(* Logix 5000 project; controller MV vendor 1 type 14 code 217 rev 31.11; software revision 31.00 *) (continued)
   MC_CH1_Log_ID : DINT := 56;
   MC_CH1_OneShot : BOOL;
   MC_CH1_PR1 : PlantItem := (CW := 2#0000_0000_0000_0000_0000_0000_0001_0000, CheckTime := 8, CheckTimer := 8);   // CH1_PR1
   MC_CH1_PR1_ALARM : ALARM_DIGITAL;
   MC_CH1_PR1_C : ALIAS FOR RIO_Rack_2:6:I.Data.6;
   MC_CH1_PR1_DR : ALIAS FOR RIO_Rack_2:5:O.Data.18;
   MC_CH1_PR1_O : ALIAS FOR RIO_Rack_2:6:I.Data.2;
   MC_CH1_PTX_AI : PlantItem := (CW := 2#0000_0000_0000_0000_1000_0000_0000_0000, CheckTime := 15, CheckTimer := 15, Scaled := 55.846878, RawInput := 9957.0);   // CH1_PTX
   MC_CH1_PTX_AI_RawInput : ALIAS FOR RIO_Rack_2:1:I.Ch6Data;   // Real Analog Input , Do Not Use In Code
   MC_CH1_R1 : PlantItem := (CW := 2#0000_0000_0000_0000_0000_0000_0011_0000, CheckTime := 20, CheckTimer := 20);   // CH1_R1
   MC_CH1_R1_ALARM : ALARM_DIGITAL;
   MC_CH1_R1_C : ALIAS FOR RIO_Rack_2:4:I.Data.4;
   MC_CH1_R1_DR : ALIAS FOR RIO_Rack_2:5:O.Data.0;
   MC_CH1_R1_O : ALIAS FOR RIO_Rack_2:4:I.Data.0;
   MC_CH1_R1R : PlantItem := (CW := 2#0000_0000_0000_0000_0000_0000_0001_0000, CheckTime := 20, CheckTimer := 20);   // CH1_R1R
   MC_CH1_R1R_ALARM : ALARM_DIGITAL;
   MC_CH1_R1R_C : ALIAS FOR RIO_Rack_2:4:I.Data.14;
   MC_CH1_R1R_DR : ALIAS FOR RIO_Rack_2:5:O.Data.6;
   MC_CH1_R1R_O : ALIAS FOR RIO_Rack_2:4:I.Data.10;
   MC_CH1_R2 : PlantItem := (CW := 2#0000_0000_0000_0000_0000_0000_0001_0000, CheckTime := 20, CheckTimer := 20);   // CH1_R2
   MC_CH1_R2_ALARM : ALARM_DIGITAL;
   MC_CH1_R2_C : ALIAS FOR RIO_Rack_2:4:I.Data.5;
   MC_CH1_R2_DR : ALIAS FOR RIO_Rack_2:5:O.Data.1;
   MC_CH1_R2_O : ALIAS FOR RIO_Rack_2:4:I.Data.1;
   MC_CH1_R2R : PlantItem := (CW := 2#0000_0000_0000_0000_0000_0000_0001_0000, CheckTime := 20, CheckTimer := 20);   // CH1_R2R
   MC_CH1_R2R_ALARM : ALARM_DIGITAL;
   MC_CH1_R2R_C : ALIAS FOR RIO_Rack_2:4:I.Data.15;
   MC_CH1_R2R_DR : ALIAS FOR RIO_Rack_2:5:O.Data.7;
   MC_CH1_R2R_O : ALIAS FOR RIO_Rack_2:4:I.Data.11;
   MC_CH1_R3 : PlantItem := (CW := 2#0000_0000_0000_0000_0000_0000_0001_0000, CheckTime := 20, CheckTimer := 20);   // CH1_R3
   MC_CH1_R3_ALARM : ALARM_DIGITAL;
   MC_CH1_R3_C : ALIAS FOR RIO_Rack_2:4:I.Data.6;
   MC_CH1_R3_DR : ALIAS FOR RIO_Rack_2:5:O.Data.2;
   MC_CH1_R3_O : ALIAS FOR RIO_Rack_2:4:I.Data.2;
   MC_CH1_R3R : PlantItem := (CW := 2#0000_0000_0000_0000_0000_0000_0001_0000, CheckTime := 20, CheckTimer := 20);   // CH1_R3R
   MC_CH1_R3R_ALARM : ALARM_DIGITAL;
   MC_CH1_R3R_C : ALIAS FOR RIO_Rack_2:4:I.Data.20;
   MC_CH1_R3R_DR : ALIAS FOR RIO_Rack_2:5:O.Data.8;
   MC_CH1_R3R_O : ALIAS FOR RIO_Rack_2:4:I.Data.16;
   MC_CH1_R4 : PlantItem := (CW := 2#0000_0000_0000_0000_0000_0000_0001_0000, CheckTime := 20, CheckTimer := 20);   // CH1_R4
   MC_CH1_R4_ALARM : ALARM_DIGITAL;
   MC_CH1_R4_C : ALIAS FOR RIO_Rack_2:4:I.Data.7;
   MC_CH1_R4_DR : ALIAS FOR RIO_Rack_2:5:O.Data.3;
   MC_CH1_R4_O : ALIAS FOR RIO_Rack_2:4:I.Data.3;
   MC_CH1_R4R : PlantItem := (CW := 2#0000_0000_0000_0000_0000_0000_0001_0000, CheckTime := 20, CheckTimer := 20);   // CH1_R4R
   MC_CH1_R4R_ALARM : ALARM_DIGITAL;
   MC_CH1_R4R_C : ALIAS FOR RIO_Rack_2:4:I.Data.21;
   MC_CH1_R4R_DR : ALIAS FOR RIO_Rack_2:5:O.Data.9;
   MC_CH1_R4R_O : ALIAS FOR RIO_Rack_2:4:I.Data.17;
   MC_CH1_R5 : PlantItem := (CW := 2#0000_0000_0000_0000_0000_0000_0001_0000, CheckTime := 20, CheckTimer := 20);   // CH1_R5
   MC_CH1_R5_ALARM : ALARM_DIGITAL;
   MC_CH1_R5_C : ALIAS FOR RIO_Rack_2:4:I.Data.12;
   MC_CH1_R5_DR : ALIAS FOR RIO_Rack_2:5:O.Data.4;
   MC_CH1_R5_O : ALIAS FOR RIO_Rack_2:4:I.Data.8;
   MC_CH1_R5R : PlantItem := (CW := 2#0000_0000_0000_0000_0000_0000_0001_0000, CheckTime := 20, CheckTimer := 20);   // CH1_R5R
   MC_CH1_R5R_ALARM : ALARM_DIGITAL;
   MC_CH1_R5R_C : ALIAS FOR RIO_Rack_2:4:I.Data.22;
   MC_CH1_R5R_DR : ALIAS FOR RIO_Rack_2:5:O.Data.10;
   MC_CH1_R5R_O : ALIAS FOR RIO_Rack_2:4:I.Data.18;
   MC_CH1_R6 : PlantItem := (CW := 2#0000_0000_0000_0000_0000_0000_1000_1011, CheckTime := 20, CheckTimer := 20, DriveBits := 1);   // CH1_R6
   MC_CH1_R6_ALARM : ALARM_DIGITAL;
   MC_CH1_R6_C : ALIAS FOR RIO_Rack_2:4:I.Data.13;
   MC_CH1_R6_DR : ALIAS FOR RIO_Rack_2:5:O.Data.5;
   MC_CH1_R6_O : ALIAS FOR RIO_Rack_2:4:I.Data.9;
   MC_CH1_R6R : PlantItem := (CW := 2#0000_0000_0000_0000_0000_0000_1000_1011, CheckTime := 20, CheckTimer := 20, DriveBits := 1);   // CH1_R6R
   MC_CH1_R6R_ALARM : ALARM_DIGITAL;
   MC_CH1_R6R_C : ALIAS FOR RIO_Rack_2:4:I.Data.23;
   MC_CH1_R6R_DR : ALIAS FOR RIO_Rack_2:5:O.Data.11;
   MC_CH1_R6R_O : ALIAS FOR RIO_Rack_2:4:I.Data.19;
   MC_CH1_RESET : ALIAS FOR MC_N100[30].0;   // CH1 reset flag
   MC_CH1_RESTART : ALIAS FOR MC_N100[35];   // CH1 restart step
   MC_CH1_RETURN : ALIAS FOR MC_N100[32].7;   // CH1 open return route flag
   MC_CH1_RP_OFF : ALIAS FOR MC_N100[32].2;   // CH1 enable return pump off delay timer
   MC_CH1_RP_ON : ALIAS FOR MC_N100[32].1;   // CH1 enable return pump on delay timer
   MC_CH1_RPUMP : ALIAS FOR MC_N100[32].4;   // CH1 run return pump flag
   MC_CH1_RR : PlantItem := (CW := 2#0000_0000_0000_0000_0000_0000_0001_0000, CheckTime := 20, CheckTimer := 20);   // CH1_RR
   MC_CH1_RR_ALARM : ALARM_DIGITAL;
   MC_CH1_RR_C : ALIAS FOR RIO_Rack_2:4:I.Data.29;
   MC_CH1_RR_DR : ALIAS FOR RIO_Rack_2:5:O.Data.13;
   MC_CH1_RR_O : ALIAS FOR RIO_Rack_2:4:I.Data.25;
   MC_CH1_RTNFLOW : ALIAS FOR MC_N100[18].0;   // CH1 Is Return Flow flag
   MC_CH1_SaveCIPReport_now : DINT;
   MC_CH1_SaveCIPReport_now_done : DINT := -1;
   MC_CH1_STATUS : ALIAS FOR MC_N100[0];   // CH1 status 0: Unavailable; 1: Idle; 2: Running; 3: Stopped; 4: Faulted
   MC_CH1_SUBSTEP : ALIAS FOR MC_N100[17];   // CH1 current substep
   MC_CH1_SUPPLY : ALIAS FOR MC_N100[32].3;   // CH1 open supply route flag
   MC_CH1_T105_2_ACC : DINT := 86383;
   MC_CH1_TIMING : ALIAS FOR MC_N100[30].3;   // CH1 run current cycle timer
   MC_CH1_TODET : ALIAS FOR MC_N100[18].2;   // CH1 return postrinse to detergent tank
   MC_CH2_ACTIVE : ALIAS FOR MC_N120[30].1;   // CH2 active flag
   MC_CH2_CIP_BYPASS_Conditions : BOOL;
   MC_CH2_CIP_BYPASS_DrainConditions : BOOL;
   MC_CH2_CIP_Messages : STRING[20];   // CH2 CIP Scada Messages
        [4]   // Channel 2 CIP Completion Clock Time
        [0]   // Channel 2 CIP Program Text for Scada
        [1]   // Channel2 CIP Cycle Text for Scada
        [2]   // Channel 2 CIP Time Left Text for Scada
        [3]   // Channel 2 CIP Down Time Text for Scada
   MC_CH2_CIP_Misc : DINT[20];
   MC_CH2_CIP_MiscReal : REAL[20];
   MC_CH2_CIP_YST_Scb_Bypass : BOOL;
   MC_CH2_CSTEP : ALIAS FOR MC_N120[34];   // CH2 command processor current step
   MC_CH2_CTX2_AI : PlantItem := (CW := 2#0000_0000_0000_0000_1000_0000_0000_0000, CheckTime := 15, CheckTimer := 15, Scaled := 0.00875, RawInput := 4014.0);   // CH2_CTX2
   MC_CH2_CTX2_AI_RawInput : ALIAS FOR RIO_Rack_2:1:I.Ch3Data;   // Real Analog Input , Do Not Use In Code
   MC_CH2_CYCDONE : ALIAS FOR MC_T125[2].DN;   // CH2 current cycle complete
   MC_CH2_CYCLE : ALIAS FOR MC_N120[1];   // CH2 current CIP cycle
   MC_CH2_Delay_For_Data : TIMER := (PRE := 2000);
   MC_CH2_DETRTN : ALIAS FOR MC_N120[18].1;   // CH2 Is Detergent Return flag
   MC_CH2_DONE : ALIAS FOR MC_N120[30].4;   // CH2 cycle complete flag
   MC_CH2_DR1 : PlantItem := (CW := 2#0000_0000_0000_0000_0000_0000_0001_0000, CheckTime := 8, CheckTimer := 8);   // CH2_DR1
   MC_CH2_DR1_ALARM : ALARM_DIGITAL;
   MC_CH2_DR1_C : ALIAS FOR RIO_Rack_2:7:I.Data.6;
   MC_CH2_DR1_DR : ALIAS FOR RIO_Rack_2:8:O.Data.2;
   MC_CH2_DR1_O : ALIAS FOR RIO_Rack_2:7:I.Data.2;
   MC_CH2_DR2 : PlantItem := (CW := 2#0000_0000_0000_0000_0000_0000_0001_0000, CheckTime := 8, CheckTimer := 8);   // CH2_DR2
   MC_CH2_DR2_ALARM : ALARM_DIGITAL;
   MC_CH2_DR2_C : ALIAS FOR RIO_Rack_2:7:I.Data.7;
   MC_CH2_DR2_DR : ALIAS FOR RIO_Rack_2:8:O.Data.3;
   MC_CH2_DR2_O : ALIAS FOR RIO_Rack_2:7:I.Data.3;
   MC_CH2_DRAIN : PlantItem := (CW := 2#0000_0000_0000_0000_0000_0000_0001_0000, CheckTime := 8, CheckTimer := 8);   // CH2_DRAIN
   MC_CH2_DRAIN_ALARM : ALARM_DIGITAL;
   MC_CH2_DRAIN_C : ALIAS FOR RIO_Rack_2:7:I.Data.4;
   MC_CH2_DRAIN_CLOSE : BOOL;
   MC_CH2_DRAIN_DR : ALIAS FOR RIO_Rack_2:8:O.Data.0;
   MC_CH2_DRAIN_O : ALIAS FOR RIO_Rack_2:7:I.Data.0;
   MC_CH2_DT : ALIAS FOR MC_N120[10];   // CH2 detergent tank to use (1 or 2)
   MC_CH2_DT1 : PlantItem := (CW := 2#0000_0000_0000_0000_0000_0000_0001_0000, CheckTime := 8, CheckTimer := 8);   // CH2_DT1
   MC_CH2_DT1_ALARM : ALARM_DIGITAL;
   MC_CH2_DT1_C : ALIAS FOR RIO_Rack_2:7:I.Data.12;
   MC_CH2_DT1_DR : ALIAS FOR RIO_Rack_2:8:O.Data.4;
   MC_CH2_DT1_O : ALIAS FOR RIO_Rack_2:7:I.Data.8;
   MC_CH2_DT2 : PlantItem := (CW := 2#0000_0000_0000_0000_0000_0000_0001_0000, CheckTime := 12, CheckTimer := 12);   // CH2_DT2
   MC_CH2_DT2_ALARM : ALARM_DIGITAL;
   MC_CH2_DT2_C : ALIAS FOR RIO_Rack_2:7:I.Data.13;
   MC_CH2_DT2_DR : ALIAS FOR RIO_Rack_2:8:O.Data.5;
   MC_CH2_DT2_O : ALIAS FOR RIO_Rack_2:7:I.Data.9;
   MC_CH2_EVENT : ALIAS FOR MC_N120[23];   // CH2 event register
   MC_CH2_EXTEND : ALIAS FOR MC_N120[30].5;   // CH2 extend cycle flag
   MC_CH2_FAULT : ALIAS FOR MC_N120[20];   // CH2 fault register
   MC_CH2_FM_AI : PlantItem := (CW := 2#0000_0000_0000_0000_1000_0000_0000_0000, CheckTime := 15, CheckTimer := 15, Scaled := 1.0, RawInput := 4032.0);   // CH2_FM
   MC_CH2_FM_AI_RawInput : ALIAS FOR RIO_Rack_2:1:I.Ch5Data;   // Real Analog Input , Do Not Use In Code
   MC_CH2_FVBypass_Flush_ALARM : ALARM_DIGITAL;
   MC_CH2_FVBYPASS_H2O_Flush : BOOL;
   MC_CH2_ISLINE : ALIAS FOR MC_N122[13].0;   // CH2 Is Line Clean flag
   MC_CH2_LF1 : PlantItem := (CW := 2#0000_0000_0000_0000_0000_0000_0001_0000, CheckTime := 8, CheckTimer := 8);   // CH2_LF1
   MC_CH2_LF1_ALARM : ALARM_DIGITAL;
   MC_CH2_LF1_C : ALIAS FOR RIO_Rack_2:7:I.Data.15;
   MC_CH2_LF1_DR : ALIAS FOR RIO_Rack_2:8:O.Data.7;
   MC_CH2_LF1_O : ALIAS FOR RIO_Rack_2:7:I.Data.11;
   MC_CH2_Log_ID : DINT := 57;
   MC_CH2_OneShot : BOOL;
   MC_CH2_PR1 : PlantItem := (CW := 2#0000_0000_0000_0000_0000_0000_0001_0000, CheckTime := 8, CheckTimer := 8);   // CH2_PR1
   MC_CH2_PR1_ALARM : ALARM_DIGITAL;
   MC_CH2_PR1_C : ALIAS FOR RIO_Rack_2:7:I.Data.14;
   MC_CH2_PR1_DR : ALIAS FOR RIO_Rack_2:8:O.Data.6;
   MC_CH2_PR1_O : ALIAS FOR RIO_Rack_2:7:I.Data.10;
   MC_CH2_PTX_AI : PlantItem := (CW := 2#0000_0000_0000_0000_1000_0000_0000_0000, CheckTime := 15, CheckTimer := 15, Scaled := 8.446876, RawInput := 4901.0);   // CH2_PTX
   MC_CH2_PTX_AI_RawInput : ALIAS FOR RIO_Rack_2:1:I.Ch7Data;   // Real Analog Input , Do Not Use In Code
   MC_CH2_R1 : PlantItem := (CW := 2#0000_0000_0000_0000_0000_0000_0001_0000, CheckTime := 8, CheckTimer := 8);   // CH2_R1
   MC_CH2_R1_ALARM : ALARM_DIGITAL;
   MC_CH2_R1_C : ALIAS FOR RIO_Rack_2:6:I.Data.12;
   MC_CH2_R1_DR : ALIAS FOR RIO_Rack_2:5:O.Data.20;
   MC_CH2_R1_O : ALIAS FOR RIO_Rack_2:6:I.Data.8;
   MC_CH2_R1R : PlantItem := (CW := 2#0000_0000_0000_0000_0000_0000_0001_0000, CheckTime := 8, CheckTimer := 8);   // CH2_R1R
   MC_CH2_R1R_ALARM : ALARM_DIGITAL;
   MC_CH2_R1R_C : ALIAS FOR RIO_Rack_2:6:I.Data.22;
   MC_CH2_R1R_DR : ALIAS FOR RIO_Rack_2:5:O.Data.26;
   MC_CH2_R1R_O : ALIAS FOR RIO_Rack_2:6:I.Data.18;
   MC_CH2_R2 : PlantItem := (CW := 2#0000_0000_0000_0000_0000_0000_0001_0000, CheckTime := 8, CheckTimer := 8);   // CH2_R2
   MC_CH2_R2_ALARM : ALARM_DIGITAL;
   MC_CH2_R2_C : ALIAS FOR RIO_Rack_2:6:I.Data.13;
   MC_CH2_R2_DR : ALIAS FOR RIO_Rack_2:5:O.Data.21;
   MC_CH2_R2_O : ALIAS FOR RIO_Rack_2:6:I.Data.9;
   MC_CH2_R2R : PlantItem := (CW := 2#0000_0000_0000_0000_0000_0000_0001_0000, CheckTime := 8, CheckTimer := 8);   // CH2_R2R
   MC_CH2_R2R_ALARM : ALARM_DIGITAL;
   MC_CH2_R2R_C : ALIAS FOR RIO_Rack_2:6:I.Data.23;
   MC_CH2_R2R_DR : ALIAS FOR RIO_Rack_2:5:O.Data.27;
   MC_CH2_R2R_O : ALIAS FOR RIO_Rack_2:6:I.Data.19;
   MC_CH2_R3 : PlantItem := (CW := 2#0000_0000_0000_0000_0000_0000_0001_0000, CheckTime := 8, CheckTimer := 8);   // CH2_R3
   MC_CH2_R3_ALARM : ALARM_DIGITAL;
   MC_CH2_R3_C : ALIAS FOR RIO_Rack_2:6:I.Data.14;
   MC_CH2_R3_DR : ALIAS FOR RIO_Rack_2:5:O.Data.22;
   MC_CH2_R3_O : ALIAS FOR RIO_Rack_2:6:I.Data.10;
   MC_CH2_R3R : PlantItem := (CW := 2#0000_0000_0000_0000_0000_0000_0001_0000, CheckTime := 8, CheckTimer := 8);   // CH2_R3R
   MC_CH2_R3R_ALARM : ALARM_DIGITAL;
   MC_CH2_R3R_C : ALIAS FOR RIO_Rack_2:6:I.Data.28;
   MC_CH2_R3R_DR : ALIAS FOR RIO_Rack_2:5:O.Data.28;
   MC_CH2_R3R_O : ALIAS FOR RIO_Rack_2:6:I.Data.24;
   MC_CH2_R4 : PlantItem := (CW := 2#0000_0000_0000_0000_0000_0000_0001_0000, CheckTime := 8, CheckTimer := 8);   // CH2_R4
   MC_CH2_R4_ALARM : ALARM_DIGITAL;
   MC_CH2_R4_C : ALIAS FOR RIO_Rack_2:6:I.Data.15;
   MC_CH2_R4_DR : ALIAS FOR RIO_Rack_2:5:O.Data.23;
   MC_CH2_R4_O : ALIAS FOR RIO_Rack_2:6:I.Data.11;
   MC_CH2_R4R : PlantItem := (CW := 2#0000_0000_0000_0000_0000_0000_0001_0000, CheckTime := 8, CheckTimer := 8);   // CH2_R4R
   MC_CH2_R4R_ALARM : ALARM_DIGITAL;
   MC_CH2_R4R_C : ALIAS FOR RIO_Rack_2:6:I.Data.29;
   MC_CH2_R4R_DR : ALIAS FOR RIO_Rack_2:5:O.Data.29;
   MC_CH2_R4R_O : ALIAS FOR RIO_Rack_2:6:I.Data.25;
   MC_CH2_R5 : PlantItem := (CW := 2#0000_0000_0000_0000_0000_0000_0001_0000, CheckTime := 8, CheckTimer := 8);   // CH2_R5
   MC_CH2_R5_ALARM : ALARM_DIGITAL;
   MC_CH2_R5_C : ALIAS FOR RIO_Rack_2:6:I.Data.20;
   MC_CH2_R5_DR : ALIAS FOR RIO_Rack_2:5:O.Data.24;
   MC_CH2_R5_O : ALIAS FOR RIO_Rack_2:6:I.Data.16;
   MC_CH2_R5R : PlantItem := (CW := 2#0000_0000_0000_0000_0000_0000_0001_0000, CheckTime := 8, CheckTimer := 8);   // CH2_R5R
   MC_CH2_R5R_ALARM : ALARM_DIGITAL;
   MC_CH2_R5R_C : ALIAS FOR RIO_Rack_2:6:I.Data.30;
   MC_CH2_R5R_DR : ALIAS FOR RIO_Rack_2:5:O.Data.30;
   MC_CH2_R5R_O : ALIAS FOR RIO_Rack_2:6:I.Data.26;
   MC_CH2_R6 : PlantItem := (CW := 2#0000_0000_0000_0000_0000_0001_0001_0000, CheckTime := 8, CheckTimer := 8);   // CH2_R6
   MC_CH2_R6_ALARM : ALARM_DIGITAL;
   MC_CH2_R6_C : ALIAS FOR RIO_Rack_2:6:I.Data.21;
   MC_CH2_R6_DR : ALIAS FOR RIO_Rack_2:5:O.Data.25;
   MC_CH2_R6_O : ALIAS FOR RIO_Rack_2:6:I.Data.17;
   MC_CH2_R6R : PlantItem := (CW := 2#0000_0000_0000_0000_0000_0000_0001_0000, CheckTime := 8, CheckTimer := 8);   // CH2_R6R
   MC_CH2_R6R_ALARM : ALARM_DIGITAL;
   MC_CH2_R6R_C : ALIAS FOR RIO_Rack_2:6:I.Data.31;
   MC_CH2_R6R_DR : ALIAS FOR RIO_Rack_2:5:O.Data.31;
   MC_CH2_R6R_O : ALIAS FOR RIO_Rack_2:6:I.Data.27;
   MC_CH2_RESET : ALIAS FOR MC_N120[30].0;   // CH2 reset flag
   MC_CH2_RESTART : ALIAS FOR MC_N120[35];   // CH2 restart step
   MC_CH2_RETURN : ALIAS FOR MC_N120[32].7;   // CH2 open return route flag
   MC_CH2_RP_ON : ALIAS FOR MC_N120[32].1;   // CH2 enable return pump on delay timer
   MC_CH2_RPUMP : ALIAS FOR MC_N120[32].4;   // CH2 run return pump flag
   MC_CH2_RR : PlantItem := (CW := 2#0000_0000_0000_0000_0000_0000_0001_0000, CheckTime := 8, CheckTimer := 8);   // CH2_RR
   MC_CH2_RR_ALARM : ALARM_DIGITAL;
   MC_CH2_RR_C : ALIAS FOR RIO_Rack_2:7:I.Data.5;
   MC_CH2_RR_DR : ALIAS FOR RIO_Rack_2:8:O.Data.1;
   MC_CH2_RR_O : ALIAS FOR RIO_Rack_2:7:I.Data.1;
   MC_CH2_RTNFLOW : ALIAS FOR MC_N120[18].0;   // CH2 return flow on debounce timer
   MC_CH2_SaveCIPReport_now : DINT;
   MC_CH2_SaveCIPReport_now_done : DINT := -1;
   MC_CH2_STATUS : ALIAS FOR MC_N120[0];   // CH2 status 0: Unavailable; 1: Idle; 2: Running; 3: Stopped; 4: Faulted
   MC_CH2_SUBSTEP : ALIAS FOR MC_N120[17];   // CH2 current substep
   MC_CH2_SUPPLY : ALIAS FOR MC_N120[32].3;   // CH2 open supply route flag
   MC_CH2_T125_2_ACC : DINT := 90000;
   MC_CH2_TIMING : ALIAS FOR MC_N120[30].3;   // CH2 run current cycle timer
   MC_CH2_TODET : ALIAS FOR MC_N120[18].2;   // CH2 return postrinse to detergent tank
   MC_CH2_TURBID_High : BOOL;
   MC_Channel1_Channel_1_event : STRING;
   MC_Channel1_Channel_1_event_prefix : STRING;
   MC_Channel1_Channel_2_event : STRING;
   MC_Channel1_Channel_2_event_prefix : STRING;
   MC_CIP_AV01 : PlantItem := (CW := 2#0000_0000_0000_0000_0000_0000_1000_1011, CheckTime := 8, CheckTimer := 8, DriveBits := 1);   // CIP_AV01
   MC_CIP_AV01_ALARM : ALARM_DIGITAL;
   MC_CIP_AV01_C : ALIAS FOR RIO_Rack_2:9:I.Data.23;
   MC_CIP_AV01_DR : ALIAS FOR CIP_AV01_DUMMY_DR;
   MC_CIP_AV01_O : ALIAS FOR RIO_Rack_2:9:I.Data.19;
   MC_CIP_AV02 : PlantItem := (CW := 2#0000_0000_0000_0000_0000_0000_0001_0000, CheckTime := 8, CheckTimer := 8);   // CIP_AV02
   MC_CIP_AV02_ALARM : ALARM_DIGITAL;
   MC_CIP_AV02_C : ALIAS FOR RIO_Rack_2:9:I.Data.28;
   MC_CIP_AV02_DR : ALIAS FOR RIO_Rack_2:8:O.Data.27;   // Used As Output Share Item Rung 20
   MC_CIP_AV02_O : ALIAS FOR RIO_Rack_2:9:I.Data.24;
   MC_CIP_AV05 : PlantItem := (CW := 2#0000_0000_0000_0000_0000_0000_1000_1011, CheckTime := 8, CheckTimer := 8, DriveBits := 1);   // CIP_AV05
   MC_CIP_AV05_ALARM : ALARM_DIGITAL;
   MC_CIP_AV05_C : ALIAS FOR RIO_Rack_2:9:I.Data.29;
   MC_CIP_AV05_DR : ALIAS FOR CIP_AV05_DUMMY_DR;
   MC_CIP_AV05_O : ALIAS FOR RIO_Rack_2:9:I.Data.25;
   MC_CIP_AV06 : PlantItem := (CW := 2#0000_0000_0000_0000_0000_0000_0001_0000, CheckTime := 8, CheckTimer := 8);   // CIP_AV06
   MC_CIP_AV06_ALARM : ALARM_DIGITAL;
   MC_CIP_AV06_C : ALIAS FOR RIO_Rack_2:9:I.Data.30;
   MC_CIP_AV06_DR : ALIAS FOR RIO_Rack_2:8:O.Data.28;
   MC_CIP_AV06_O : ALIAS FOR RIO_Rack_2:9:I.Data.26;
   MC_CIP_AV07 : PlantItem := (CW := 2#0000_0000_0000_0000_0000_0000_1000_1011, CheckTime := 8, CheckTimer := 8, DriveBits := 1);   // CIP_AV07
   MC_CIP_AV07_ALARM : ALARM_DIGITAL;
   MC_CIP_AV07_C : ALIAS FOR RIO_Rack_2:9:I.Data.31;
   MC_CIP_AV07_DR : ALIAS FOR CIP_AV07_DUMMY_DR;
   MC_CIP_AV07_O : ALIAS FOR RIO_Rack_2:9:I.Data.27;
   MC_CIP_AV08 : PlantItem := (CW := 2#0000_0000_0000_0000_0000_0000_0001_0000, CheckTime := 8, CheckTimer := 8);   // CIP_AV08
   MC_CIP_AV08_ALARM : ALARM_DIGITAL;
   MC_CIP_AV08_C : ALIAS FOR RIO_Rack_2:11:I.Data.20;
   MC_CIP_AV08_DR : ALIAS FOR RIO_Rack_2:8:O.Data.29;
   MC_CIP_AV08_O : ALIAS FOR RIO_Rack_2:11:I.Data.24;
   MC_CIP_AV09 : PlantItem := (CW := 2#0000_0000_0000_0000_0000_0000_1000_1011, CheckTime := 8, CheckTimer := 8, DriveBits := 1);   // CIP_AV09
   MC_CIP_AV09_ALARM : ALARM_DIGITAL;
   MC_CIP_AV09_C : ALIAS FOR RIO_Rack_2:11:I.Data.21;
   MC_CIP_AV09_DR : ALIAS FOR CIP_AV09_DUMMY_DR;
   MC_CIP_AV09_O : ALIAS FOR RIO_Rack_2:11:I.Data.25;
   MC_CIP_AV10 : PlantItem := (CW := 2#0000_0000_0000_0000_0000_0000_0001_0000, CheckTime := 8, CheckTimer := 8);   // CIP_AV10
   MC_CIP_AV10_ALARM : ALARM_DIGITAL;
   MC_CIP_AV10_C : ALIAS FOR RIO_Rack_2:11:I.Data.22;
   MC_CIP_AV10_DR : ALIAS FOR RIO_Rack_2:8:O.Data.30;
   MC_CIP_AV10_O : ALIAS FOR RIO_Rack_2:11:I.Data.26;
   MC_CIP_CH2_String_OK : BOOL;
   MC_CIP_CH2_Strings_HopRinse : STRING[30] := ([0] := 'FV', [1] := 'YSV', [2] := 'YPV', [3] := 'YCV', [4] := 'Yeast Pitch Main', [5] := 'Yeast Slurry Tank', [6] := 'Gales Yeast Main', [7] := 'YSV1 Reseeding Line', [8] := 'Filtrate Tank', [9] := 'Yeast Main FVs1 to 17 Short', [10] := 'Yeast Main FVs1 to 17 Long', [11] := 'Yeast Main FVs18 to 25 Short', [12] := 'Yeast Main FVs18 to 25 Long', [13] := 'Yeast Room and Pump', [14] := 'FVs 26 to 31 Yeast Main Short', [15] := 'FVs 26 to 31 Yeast Main Long', [16] := ' Normal Clean', [17] := ' Hop Rinse', [18] := ' Hop Normal clean 3 pre rinses', [19] := ' Initial rinse', [20] := ' Pre-CIP Initial Rinse', [21] := ' Normal', [22] := 'Cold Water Rinse');
   MC_CIP_Default_Messages : STRING[20] := ([1] := 'Scavenge ', [2] := 'Pre Rinse ', [3] := 'Detergent ', [4] := 'Post Rinse ', [5] := ' of ', [6] := ':', [7] := '0', [17] := '3', [18] := '16', [19] := '1');
        [5]   // cycle of with spaces
        [6]   // colon : for time
        [17]   // Temp Working Area
        [18]   // Temp Working Area
        [0]   // temp area to build
        [19]   // Temp Working Area
        [7]   // leading 'zero'
   MC_CIP_EFFTank_Full : BOOL;
   MC_CIP_EFFTank_Full_Spt : DINT := 50000;
   MC_CIP_EFFTank_Start_Lvl_Ok : BOOL := 1;
   MC_CIP_RV : PlantItem := (CW := 2#0000_0000_0000_0000_0000_0001_0000_0000, CheckTime := 15, CheckTimer := 15);   // CIP_RV
   MC_CIP_RV_ALARM : ALARM_DIGITAL;
   MC_CIP_RV_C : ALIAS FOR RIO_Rack_2:9:I.Data.21;
   MC_CIP_RV_DR : ALIAS FOR RIO_Rack_2:8:O.Data.26;
   MC_CIP_RV_O : ALIAS FOR RIO_Rack_2:9:I.Data.17;
   MC_CIP_String_Result : DINT;
   MC_CIP_temp : INT;
   MC_CLOCK_system_set : BOOL;
   MC_COMMS_FROM_BLUNGER : MESSAGE;
        MessageParameters(ServiceCode := 16#0fa2, LocalElement := MC_N114[0], ...)
   mc_comms_from_brewhouse : MESSAGE;
        MessageParameters(ServiceCode := 16#004c, LocalElement := BH_Draindown_ON, ...)
   mc_comms_from_brewhouse_timer : TIMER := (PRE := 6000, ACC := 1632, EN := 1, TT := 1);
   MC_COMMS_FROM_FV_ROUTING_PLC : MESSAGE;
        MessageParameters(ServiceCode := 16#004c, LocalElement := MC_N112[0], ...)
   MC_COMMS_FROM_MV_ROUTING_PLC : MESSAGE;
        MessageParameters(ServiceCode := 16#004c, LocalElement := MC_N113[0], ...)
   mc_comms_to_blunger : MESSAGE;
        MessageParameters(ServiceCode := 16#0faa, LocalElement := MC_N114[100], ...)
   mc_comms_to_blunger_timer : TIMER := (PRE := 6000, ACC := 631, EN := 1, TT := 1);
   mc_comms_to_fv_route : MESSAGE;
        MessageParameters(ServiceCode := 16#0faa, LocalElement := MC_N112[100], ...)
   mc_comms_to_fv_route_timer : TIMER := (PRE := 6000, ACC := 2121, EN := 1, TT := 1);
   mc_comms_to_mv_route : MESSAGE;
        MessageParameters(ServiceCode := 16#0faa, LocalElement := MC_N113[100], ...)
   mc_comms_to_mv_route_timer : TIMER := (PRE := 6000, ACC := 629, EN := 1, TT := 1);
   MC_copy_how_many : DINT;
   MC_CopyOfCh1Route : DINT := 1032;
   MC_CopyOfCh2Route : DINT := 7;
   MC_CP1 : PlantItem := (CheckTime := 8);   // CP1
   MC_CP1_RawOutput : ALIAS FOR RIO_Rack_2:10:O.Data.14;   // MC_CP1
   MC_CTX_001_AI : PlantItem := (CW := 2#0000_0000_0000_0000_1100_0000_0000_0000, CheckTime := 15, CheckTimer := 15, Scaled := 2.2806249, RawInput := 7649.0);   // CTX_001
   MC_CTX_001_AI_RawInput : ALIAS FOR RIO_Rack_2:1:I.Ch0Data;   // Real Analog Input , Do Not Use In Code
   MC_CTX_002_AI : PlantItem := (CW := 2#0000_0000_0000_0000_1000_0000_0000_0000, CheckTime := 15, CheckTimer := 15, Scaled := 2.170625, RawInput := 7473.0);   // CTX_002
   MC_CTX_002_AI_RawInput : ALIAS FOR RIO_Rack_2:1:I.Ch1Data;   // Real Analog Input , Do Not Use In Code
   MC_data_file_address : DINT := 80;
   MC_data_file_value_to_move : DINT := 18;
   MC_Delphi_I : DINT[60] := ([38] := 29712, [39] := 33151);
   MC_DetTank1_Service_event : STRING;
   MC_DetTank1_Service_event_prefix : STRING;
   MC_DetTank2_Service_event : STRING;
   MC_DetTank2_Service_event_prefix : STRING;
   MC_DT1_CP1 : ALIAS FOR MC_N80[18].8;   // DT1 service drive caustic pump flag
   MC_DT1_DILUTE : ALIAS FOR MC_N80[6].2;   // DT1 detergent diluted
   MC_DT1_STR_OK : ALIAS FOR MC_N80[6].0;   // DT1 detergent strength ok
   MC_DT1_TEMP_OK : ALIAS FOR MC_N80[6].1;   // DT1 detergent temperature ok
   MC_DT2_CP1 : ALIAS FOR MC_N90[18].8;   // DT2 service drive caustic pump flag
   MC_DT2_DILUTE : ALIAS FOR MC_N90[6].2;   // DT2 detergent diluted
   MC_DT2_STR_OK : ALIAS FOR MC_N90[6].0;   // DT2 detergent strength ok
   MC_DT2_TEMP_OK : ALIAS FOR MC_N90[6].1;   // DT2 detergent temperature ok
   MC_Event_Alarm_Tag : ALARM_DIGITAL;
   MC_Event_control_FIFO : CONTROL := (LEN := 30, EM := 1);
   MC_Event_control_FIFO_Operation_Type : CONTROL := (LEN := 30, EM := 1);
   MC_Event_Delay_For_Data : TIMER := (PRE := 1000);
   MC_Event_Delay_For_PLC_Startup_Data : TIMER := (PRE := 1000);
   MC_Event_Delay_Timer : TIMER := (PRE := 1000);
   MC_Event_Delay_Timer_Off : TIMER := (PRE := 1000);
   MC_Event_from_buffer : STRING := 'CIP Channel 1 Racking Main Normal clean started by operator (Amanda_H)';
   MC_Event_from_buffer_LogData1 : REAL;
   MC_Event_from_buffer_LogData2 : REAL;
   MC_Event_from_buffer_LogData3 : REAL;
   MC_Event_from_buffer_LogData4 : REAL;
   MC_Event_from_buffer_Operation_Type : DINT := 56;
   MC_event_step : DINT;
   MC_Event_String_Last : STRING := 'CIP Channel 1 Racking Main Normal clean started by operator (Amanda_H)';
   MC_Event_Transact_Trigger_Tag : DINT;
   MC_Events_FIFO_Buffer : STRING[31];
   MC_Events_FIFO_Buffer_Operation_Type : INT[31];
   MC_FL_D1 : PlantItem := (CW := 2#0000_0000_0000_0000_0000_0000_0001_0000, CheckTime := 8, CheckTimer := 8);   // FL_D1
   MC_FL_D1_ALARM : ALARM_DIGITAL;
   MC_FL_D1_C : ALIAS FOR RIO_Rack_2:7:I.Data.21;
   MC_FL_D1_DR : ALIAS FOR RIO_Rack_2:8:O.Data.9;
   MC_FL_D1_O : ALIAS FOR RIO_Rack_2:7:I.Data.17;
   MC_FL_D2 : PlantItem := (CW := 2#0000_0000_0000_0000_0000_0000_0001_0000, CheckTime := 8, CheckTimer := 8);   // FL_D2
   MC_FL_D2_ALARM : ALARM_DIGITAL;
   MC_FL_D2_C : ALIAS FOR RIO_Rack_2:7:I.Data.22;
   MC_FL_D2_DR : ALIAS FOR RIO_Rack_2:8:O.Data.10;
   MC_FL_D2_O : ALIAS FOR RIO_Rack_2:7:I.Data.18;
   MC_FL_PR : PlantItem := (CW := 2#0000_0000_0000_0000_0000_0000_0001_0000, CheckTime := 8, CheckTimer := 8);   // FL_PR
   MC_FL_PR_ALARM : ALARM_DIGITAL;
   MC_FL_PR_C : ALIAS FOR RIO_Rack_2:7:I.Data.20;
   MC_FL_PR_DR : ALIAS FOR RIO_Rack_2:8:O.Data.8;
   MC_FL_PR_O : ALIAS FOR RIO_Rack_2:7:I.Data.16;
   MC_from_data_file : DINT := 80;
   MC_from_data_offset : DINT := 21;
   MC_FVR_FAIL : ALIAS FOR MC_N112[20].0;   // Comms.to FV Routing PLC have failed
   MC_FVYST_PX1 : ALIAS FOR MC_N112[10].0;
   MC_FVYST_PX2 : ALIAS FOR MC_N112[10].1;
   MC_FVYST_PX3 : ALIAS FOR MC_N112[10].2;
   MC_GBYV1 : PlantItem := (CheckTime := 8);   // GBYV1
   MC_GBYV1_RawOutput : ALIAS FOR RIO_Rack_2:8:O.Data.31;   // MC_GBYV1
   MC_ITEMOUT_RawOutput : ALIAS FOR RIO_Rack_2:10:O.Data.14;   // MC_ITEMOUT
   MC_Last_LogData_For_Op : REAL[60,20] := ([1,1] := 402.0, [2,1] := 33.0, [2,2] := 403.0);
   MC_LTX001_1_ON : ALIAS FOR MC_T4[1].DN;   // Prerinse tank High LP covered
   MC_LTX001_2_ON : ALIAS FOR MC_T4[2].DN;   // Prerinse tank Working LP covered
   MC_LTX001_3_OFF : ALIAS FOR MC_T4[3].DN;   // Prerinse tank Low LP not covered
   MC_LTX002_1_ON : ALIAS FOR MC_T4[4].DN;   // DT1 High LP covered
   MC_LTX002_2_ON : ALIAS FOR MC_T4[5].DN;   // DT1 Working LP covered
   MC_LTX002_3_OFF : ALIAS FOR MC_T4[6].DN;   // DT1 Low LP not covered
   MC_LTX003_1_ON : ALIAS FOR MC_T4[7].DN;   // DT2 High LP covered
   MC_LTX003_2_ON : ALIAS FOR MC_T4[8].DN;   // DT2 Working LP covered
   MC_LTX003_3_OFF : ALIAS FOR MC_T4[9].DN;   // DT2 Low LP not covered
   MC_LTX_001_1 : PlantItem := (CW := 2#0000_0000_0000_0100_0000_0000_0010_0001);   // LTX_001_1
   MC_LTX_001_1_RawInput : ALIAS FOR RIO_Rack_2:12:I.Data.16;   // MC_LTX_001_1
   MC_LTX_001_2 : PlantItem := (CW := 2#0000_0000_0000_0100_0000_0000_0000_0001, DebounceTime := 5);   // LTX_001_2
   MC_LTX_001_2_RawInput : ALIAS FOR RIO_Rack_2:12:I.Data.17;   // MC_LTX_001_2
   MC_LTX_001_3 : PlantItem := (CW := 2#0000_0000_0000_0100_0000_0000_0000_0001);   // LTX_001_3
   MC_LTX_001_3_RawInput : ALIAS FOR RIO_Rack_2:12:I.Data.18;   // MC_LTX_001_3
   MC_LTX_002_1 : PlantItem := (CW := 2#0000_0000_0000_0100_0000_0000_0000_0001);   // LTX_002_1
   MC_LTX_002_1_RawInput : ALIAS FOR RIO_Rack_2:12:I.Data.19;   // MC_LTX_002_1
   MC_LTX_002_2 : PlantItem := (CW := 2#0000_0000_0000_0100_0000_0000_0000_0001, DebounceTime := 4);   // LTX_002_2
   MC_LTX_002_2_RawInput : ALIAS FOR RIO_Rack_2:12:I.Data.20;   // MC_LTX_002_2
   MC_LTX_002_3 : PlantItem := (CW := 2#0000_0000_0000_0100_0000_0000_0010_0001);   // LTX_002_3
   MC_LTX_002_3_RawInput : ALIAS FOR RIO_Rack_2:12:I.Data.21;   // MC_LTX_002_3
   MC_LTX_003_1 : PlantItem := (CW := 2#0000_0000_0000_0100_0000_0000_0000_0001);   // LTX_003_1
   MC_LTX_003_1_RawInput : ALIAS FOR RIO_Rack_2:12:I.Data.22;   // MC_LTX_003_1
   MC_LTX_003_2 : PlantItem;   // LTX_003_2
   MC_LTX_003_2_RawInput : ALIAS FOR RIO_Rack_2:12:I.Data.23;   // MC_LTX_003_2
   MC_LTX_003_3 : PlantItem := (CW := 2#0000_0000_0000_0100_0000_0000_0010_0001);   // LTX_003_3
   MC_LTX_003_3_RawInput : ALIAS FOR RIO_Rack_2:12:I.Data.24;   // MC_LTX_003_3
   MC_MVR_FAIL : ALIAS FOR MC_N113[20].0;   // Comms.to MV Routing PLC have failed
   MC_N10 : INT[255] := ([2] := 450, [3] := 5, [4] := 11, [6] := 4, [7] := 3, [8] := 60, [9] := 500, [10] := 300, [11] := 60, [12] := 240, [13] := 3000, [14] := 23, [15] := 650, [16] := 7, [17] := 30, [18] := 480, [19] := 5, [20] := 300, [21] := 60, [22] := 180, [23] := 3000, [24] := 22, [25] := 650);   // SETTINGS
        [18]   // Eff Tank Level too high setpoint
        [14]   // DT1 service target detergent strength
        [24]   // DT2 service target detergent strength
        [7]   // Automatic timed service start hour
        [8]   // Automatic timed service start min.
        [0].0   // Request system settings reload from PC flag
        [12]   // DT1 service make-up timeout
        [13]   // DT1 service heat-up timeout
        [0].1   // Request time update from PC flag
        [22]   // DT2 service make-up timeout
        [23]   // DT2 service heat-up timeout
        [11]   // DT1 service recirc. time
        [21]   // DT2 service recirc. time
        [16]   // Turbidity meter setpoint
        [19]   // Turbidity debounce timer
        [15]   // DT1 service target temperature
        [25]   // DT2 service target temperature
        [9]   // Effluent Tank High Level Setpoint
        [10]   // DT1 service top-up timeout
        [17]   // FV Bypass Water Flush Timer
        [6]   // Current day of week (1-7: 1 = Sunday)
        [1].0   // PC has updated time flag
        [20]   // DT2 service top-up timeout
        [4]   // Current time hours (from PC)
        [5]   // Current time mins. (from PC)
   MC_N100 : INT[255] := ([0] := 2, [1] := 30, [2] := 164, [3] := 1, [4] := 1, [5] := 85, [6] := 16, [7] := 24, [10] := 1, [11] := 6, [12] := 17, [13] := 1017, [15] := 11068, [17] := 340, [18] := 3, [19] := 9, [20] := -1, [21] := 1, [22] := 2, [24] := 1, [25] := 2, [26] := -1, [29] := 20, [30] := 14, [31] := 1030, [32] := 392, [33] := 3, [34] := -1, [35] := 320, [38] := 80, [39] := 217);   // C1_PLC Channel 1 PLC data
        [31].2   // CH1 detergent initialised
        [18].3   // CH1 enable postrinse return to detergent tank
        [0]   // CH1 status 0: Unavailable; 1: Idle; 2: Running; 3: Stopped; 4: Faulted
        [31].3   // CH1 postrinse initialised
        [32].8   // CH1 route return to detergent tank flag
        [18].2   // CH1 return postrinse to detergent tank
        [32].2   // CH1 enable return pump off delay timer
        [30].3   // CH1 run current cycle timer
        [2].3   // Channel 1 continue button available
        [32].9   // CH1 initialise supply pump PID flag
        [18].1   // CH1 Is Detergent Return flag
        [2].6   // Channel 1 end extend available
        [6]   // CH1 current CIP total time minutes
        [7]   // CH1 current CIP total time seconds
        [12]   // CH1 current CIP program no.
        [18].0   // CH1 Is Return Flow flag
        [10]   // CH1 detergent tank to use (1 or 2)
        [19].1   // P1 PID pressure control selected
        [30].4   // CH1 cycle complete flag
        [19].3   // P1 PID flowrate control selected
        [28].0   // CH1 MV Routing PLC in use flag
        [28].1   // CH1 FV Routing PLC in use flag
        [27].3   // CH1 drive new route 3 routing valves
        [27].4   // CH1 drive new route 4 routing valves
        [27].5   // CH1 drive new route 5 routing valves
        [27].6   // CH1 drive new route 6 routing valves
        [32].6   // CH1 run detergent return check timer
        [33].0   // CH1 open detergent tank return valve
        [33].1   // CH1 open detergent tank outlet valve
        [2].0   // Channel 1 start button available
        [2].1   // CH1 startup in progress
        [30].2   // Channel 1 initialised
        [30].5   // CH1 extend cycle flag
        [31].10   // CH1 detergent active
        [31].11   // CH1 postrinse active
        [20]   // CH1 fault register
        [32].1   // CH1 enable return pump on delay timer
        [8]   // CH1 current CIP total stopped time minutes
        [9]   // CH1 current CIP total stopped time seconds
        [4]   // CH1 total subcycles to do
        [32].3   // CH1 open supply route flag
        [32].7   // CH1 open return route flag
        [23]   // CH1 event register
        [30].0   // CH1 reset flag
        [33].4   // CH1 detergent tank low level probe uncovered
        [17]   // CH1 current substep
        [19]   // CH1 PID flags /0: Press.inhibited /1: Press.selected /2: Flow inhibited /3: Flow selected
        [2].2   // Channel 1 stop button available
        [30].1   // CH1 active flag
        [2].4   // Channel 1 abort button availble
        [2].7   // Channel 1 skip button available
        [33].3   // CH1 detergent tank working level probe covered
        [1]   // CH1 current CIP cycle
        [21]   // CH1 fault parameter #1
        [22]   // CH1 fault parameter #2
        [24]   // CH1 event parameter #1
        [25]   // CH1 event parameter #2
        [31].8   // CH1 scavenge active
        [31].9   // CH1 prerinse active
        [3]   // CH1 current subcycle no.
        [18].4   // CH1 waiting for DT service flag
        [28].2   // CH1 Yeast Press PLC in use flag
        [5]   // CH1 time left this cycle